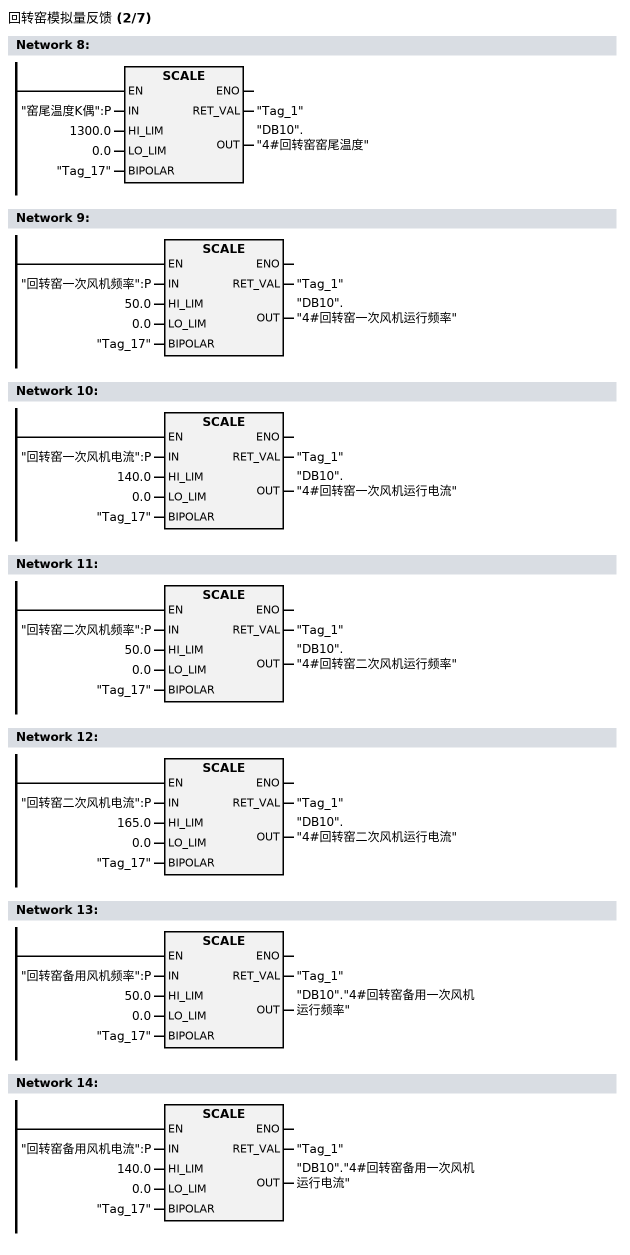
   "Tag_1" := SCALE(IN := "窑尾温度K偶":P,
                    HI_LIM := 1300.0,
                    LO_LIM := 0.0,
                    BIPOLAR := "Tag_17",
                    OUT => "DB10"."4#回转窑窑尾温度");
END_REGION

REGION Network 9
   "Tag_1" := SCALE(IN := "回转窑一次风机频率":P,
                    HI_LIM := 50.0,
                    LO_LIM := 0.0,
                    BIPOLAR := "Tag_17",
                    OUT => "DB10"."4#回转窑一次风机运行频率");
END_REGION

REGION Network 10
   "Tag_1" := SCALE(IN := "回转窑一次风机电流":P,
                    HI_LIM := 140.0,
                    LO_LIM := 0.0,
                    BIPOLAR := "Tag_17",
                    OUT => "DB10"."4#回转窑一次风机运行电流");
END_REGION

REGION Network 11
   "Tag_1" := SCALE(IN := "回转窑二次风机频率":P,
                    HI_LIM := 50.0,
                    LO_LIM := 0.0,
                    BIPOLAR := "Tag_17",
                    OUT => "DB10"."4#回转窑二次风机运行频率");
END_REGION

REGION Network 12
   "Tag_1" := SCALE(IN := "回转窑二次风机电流":P,
                    HI_LIM := 165.0,
                    LO_LIM := 0.0,
                    BIPOLAR := "Tag_17",
                    OUT => "DB10"."4#回转窑二次风机运行电流");
END_REGION

REGION Network 13
   "Tag_1" := SCALE(IN := "回转窑备用风机频率":P,
                    HI_LIM := 50.0,
                    LO_LIM := 0.0,
                    BIPOLAR := "Tag_17",
                    OUT => "DB10"."4#回转窑备用一次风机运行频率");
END_REGION

REGION Network 14
   "Tag_1" := SCALE(IN := "回转窑备用风机电流":P,
                    HI_LIM := 140.0,
                    LO_LIM := 0.0,
                    BIPOLAR := "Tag_17",
                    OUT => "DB10"."4#回转窑备用一次风机运行电流");
END_REGION

REGION Network 15
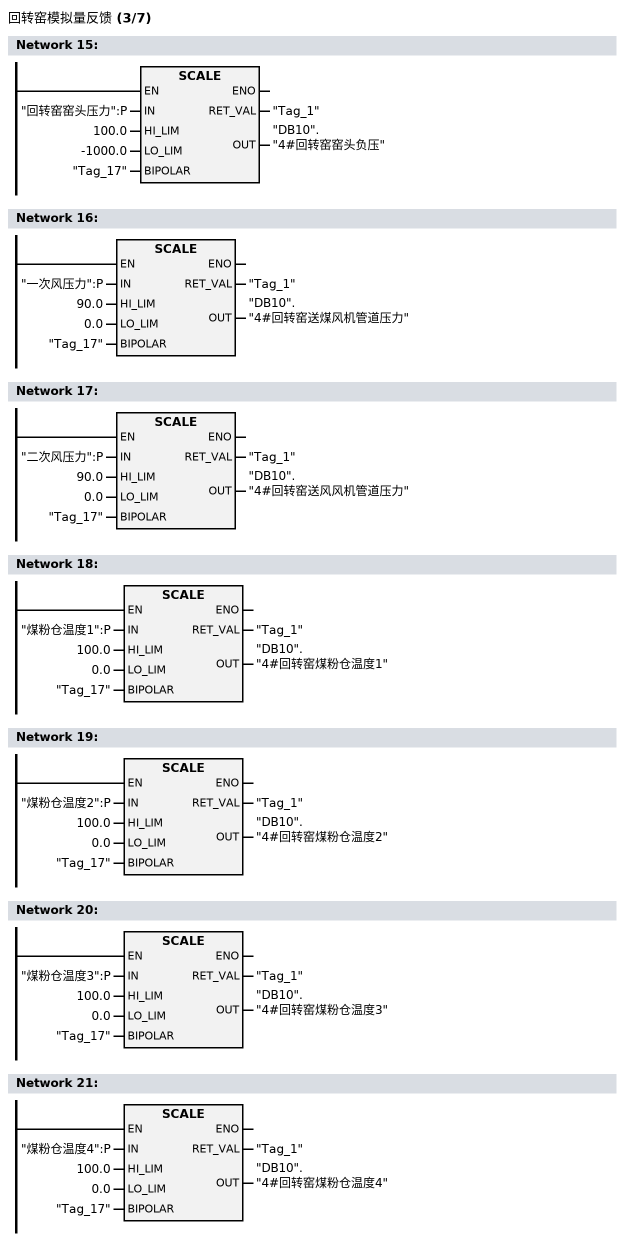
   "Tag_1" := SCALE(IN := "回转窑窑头压力":P,
                    HI_LIM := 100.0,
                    LO_LIM := -1000.0,
                    BIPOLAR := "Tag_17",
                    OUT => "DB10"."4#回转窑窑头负压");
END_REGION

REGION Network 16
   "Tag_1" := SCALE(IN := "一次风压力":P,
                    HI_LIM := 90.0,
                    LO_LIM := 0.0,
                    BIPOLAR := "Tag_17",
                    OUT => "DB10"."4#回转窑送煤风机管道压力");
END_REGION

REGION Network 17
   "Tag_1" := SCALE(IN := "二次风压力":P,
                    HI_LIM := 90.0,
                    LO_LIM := 0.0,
                    BIPOLAR := "Tag_17",
                    OUT => "DB10"."4#回转窑送风风机管道压力");
END_REGION

REGION Network 18
   "Tag_1" := SCALE(IN := "煤粉仓温度1":P,
                    HI_LIM := 100.0,
                    LO_LIM := 0.0,
                    BIPOLAR := "Tag_17",
                    OUT => "DB10"."4#回转窑煤粉仓温度1");
END_REGION

REGION Network 19
   "Tag_1" := SCALE(IN := "煤粉仓温度2":P,
                    HI_LIM := 100.0,
                    LO_LIM := 0.0,
                    BIPOLAR := "Tag_17",
                    OUT => "DB10"."4#回转窑煤粉仓温度2");
END_REGION

REGION Network 20
   "Tag_1" := SCALE(IN := "煤粉仓温度3":P,
                    HI_LIM := 100.0,
                    LO_LIM := 0.0,
                    BIPOLAR := "Tag_17",
                    OUT => "DB10"."4#回转窑煤粉仓温度3");
END_REGION

REGION Network 21
   "Tag_1" := SCALE(IN := "煤粉仓温度4":P,
                    HI_LIM := 100.0,
                    LO_LIM := 0.0,
                    BIPOLAR := "Tag_17",
                    OUT => "DB10"."4#回转窑煤粉仓温度4");
END_REGION

REGION Network 22
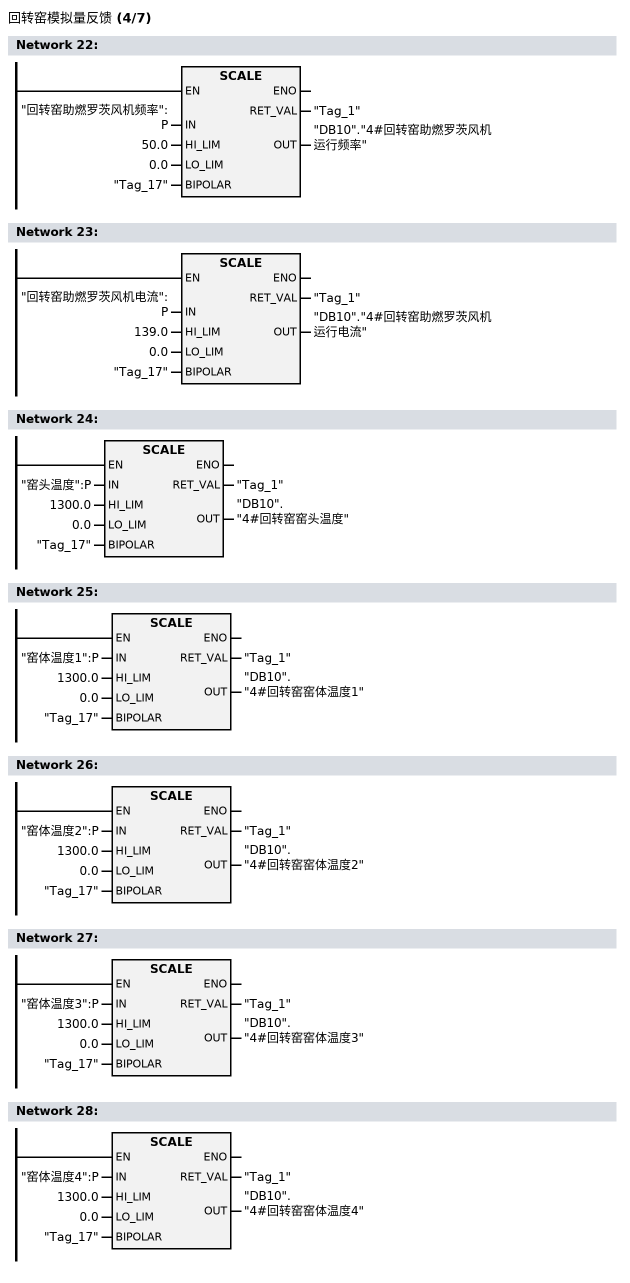
   "Tag_1" := SCALE(IN := "回转窑助燃罗茨风机频率":P,
                    HI_LIM := 50.0,
                    LO_LIM := 0.0,
                    BIPOLAR := "Tag_17",
                    OUT => "DB10"."4#回转窑助燃罗茨风机运行频率");
END_REGION

REGION Network 23
   "Tag_1" := SCALE(IN := "回转窑助燃罗茨风机电流":P,
                    HI_LIM := 139.0,
                    LO_LIM := 0.0,
                    BIPOLAR := "Tag_17",
                    OUT => "DB10"."4#回转窑助燃罗茨风机运行电流");
END_REGION

REGION Network 24
   "Tag_1" := SCALE(IN := "窑头温度":P,
                    HI_LIM := 1300.0,
                    LO_LIM := 0.0,
                    BIPOLAR := "Tag_17",
                    OUT => "DB10"."4#回转窑窑头温度");
END_REGION

REGION Network 25
   "Tag_1" := SCALE(IN := "窑体温度1":P,
                    HI_LIM := 1300.0,
                    LO_LIM := 0.0,
                    BIPOLAR := "Tag_17",
                    OUT => "DB10"."4#回转窑窑体温度1");
END_REGION

REGION Network 26
   "Tag_1" := SCALE(IN := "窑体温度2":P,
                    HI_LIM := 1300.0,
                    LO_LIM := 0.0,
                    BIPOLAR := "Tag_17",
                    OUT => "DB10"."4#回转窑窑体温度2");
END_REGION

REGION Network 27
   "Tag_1" := SCALE(IN := "窑体温度3":P,
                    HI_LIM := 1300.0,
                    LO_LIM := 0.0,
                    BIPOLAR := "Tag_17",
                    OUT => "DB10"."4#回转窑窑体温度3");
END_REGION

REGION Network 28
   "Tag_1" := SCALE(IN := "窑体温度4":P,
                    HI_LIM := 1300.0,
                    LO_LIM := 0.0,
                    BIPOLAR := "Tag_17",
                    OUT => "DB10"."4#回转窑窑体温度4");
END_REGION

REGION Network 29
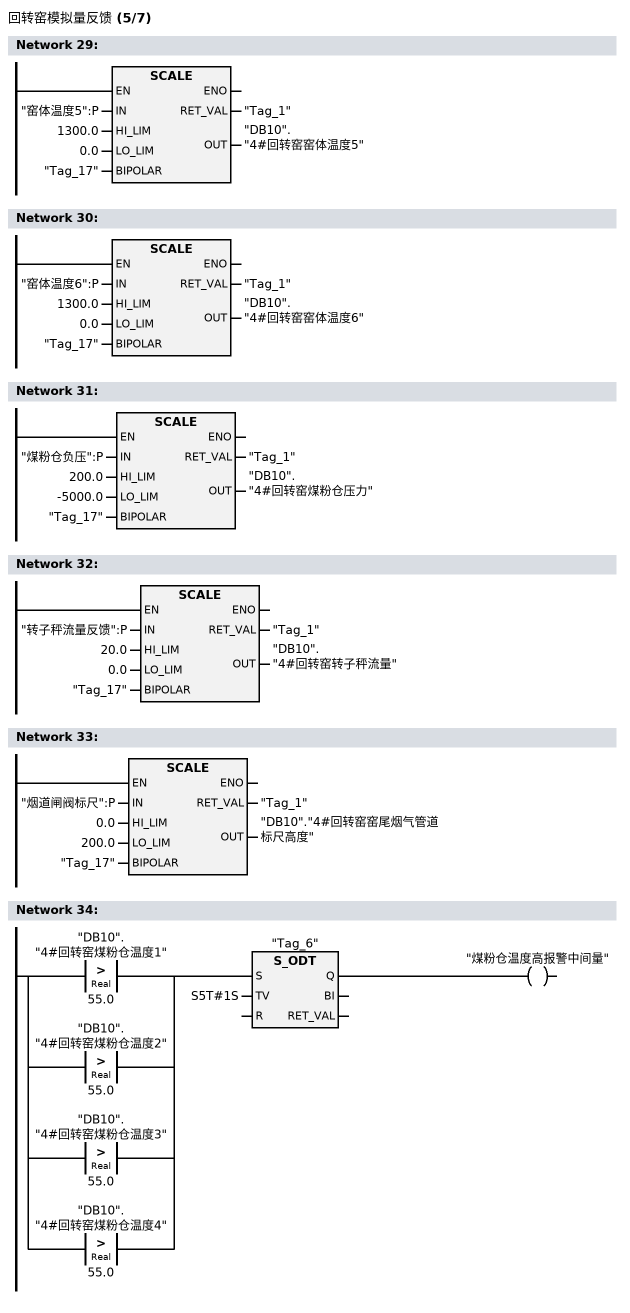
   "Tag_1" := SCALE(IN := "窑体温度5":P,
                    HI_LIM := 1300.0,
                    LO_LIM := 0.0,
                    BIPOLAR := "Tag_17",
                    OUT => "DB10"."4#回转窑窑体温度5");
END_REGION

REGION Network 30
   "Tag_1" := SCALE(IN := "窑体温度6":P,
                    HI_LIM := 1300.0,
                    LO_LIM := 0.0,
                    BIPOLAR := "Tag_17",
                    OUT => "DB10"."4#回转窑窑体温度6");
END_REGION

REGION Network 31
   "Tag_1" := SCALE(IN := "煤粉仓负压":P,
                    HI_LIM := 200.0,
                    LO_LIM := -5000.0,
                    BIPOLAR := "Tag_17",
                    OUT => "DB10"."4#回转窑煤粉仓压力");
END_REGION

REGION Network 32
   "Tag_1" := SCALE(IN := "转子秤流量反馈":P,
                    HI_LIM := 20.0,
                    LO_LIM := 0.0,
                    BIPOLAR := "Tag_17",
                    OUT => "DB10"."4#回转窑转子秤流量");
END_REGION

REGION Network 33
   "Tag_1" := SCALE(IN := "烟道闸阀标尺":P,
                    HI_LIM := 0.0,
                    LO_LIM := 200.0,
                    BIPOLAR := "Tag_17",
                    OUT => "DB10"."4#回转窑窑尾烟气管道标尺高度");
END_REGION

REGION Network 34
   RUNG wire#powerrail
      { S7_Templates := "SrcType := Real" } GT_Contact(in1 := "DB10"."4#回转窑煤粉仓温度1", in2 := 55.0)
      wire#w1
      S_ODT(T_NO := "Tag_6", TV := S5T#1S, R :=, BI =>, RET_VAL =>)
      Coil( "煤粉仓温度高报警中间量" )
   END_RUNG
   RUNG wire#powerrail
      { S7_Templates := "SrcType := Real" } GT_Contact(in1 := "DB10"."4#回转窑煤粉仓温度2", in2 := 55.0)
   END_RUNG wire#w1
   RUNG wire#powerrail
      { S7_Templates := "SrcType := Real" } GT_Contact(in1 := "DB10"."4#回转窑煤粉仓温度3", in2 := 55.0)
   END_RUNG wire#w1
   RUNG wire#powerrail
      { S7_Templates := "SrcType := Real" } GT_Contact(in1 := "DB10"."4#回转窑煤粉仓温度4", in2 := 55.0)
   END_RUNG wire#w1
   // the same network as SCL:
   #_s5time1 := S_ODT(T_NO := "Tag_6",
                      S := ("DB10"."4#回转窑煤粉仓温度1" > 55.0) OR ("DB10"."4#回转窑煤粉仓温度2" > 55.0) OR ("DB10"."4#回转窑煤粉仓温度3" > 55.0) OR ("DB10"."4#回转窑煤粉仓温度4" > 55.0),
                      TV := S5T#1S,
                      Q => #_w1);
   "煤粉仓温度高报警中间量" := #_w1;
END_REGION

REGION Network 35
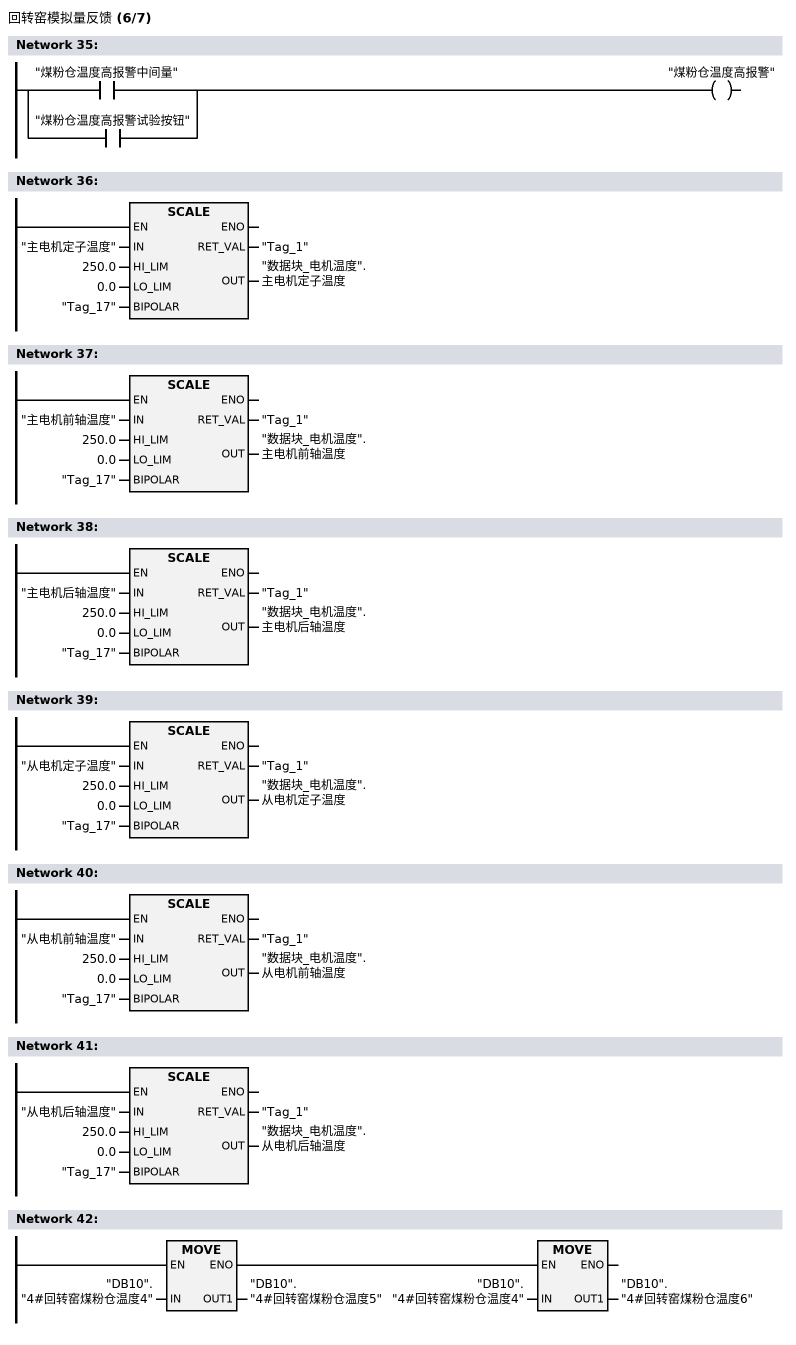
   RUNG wire#powerrail
      Contact( "煤粉仓温度高报警中间量" )
      wire#w1
      Coil( "煤粉仓温度高报警" )
   END_RUNG
   RUNG wire#powerrail
      Contact( "煤粉仓温度高报警试验按钮" )
   END_RUNG wire#w1
   // the same network as SCL:
   "煤粉仓温度高报警" := "煤粉仓温度高报警中间量" OR "煤粉仓温度高报警试验按钮";
END_REGION

REGION Network 36
   "Tag_1" := SCALE(IN := "主电机定子温度",
                    HI_LIM := 250.0,
                    LO_LIM := 0.0,
                    BIPOLAR := "Tag_17",
                    OUT => "数据块_电机温度".主电机定子温度);
END_REGION

REGION Network 37
   "Tag_1" := SCALE(IN := "主电机前轴温度",
                    HI_LIM := 250.0,
                    LO_LIM := 0.0,
                    BIPOLAR := "Tag_17",
                    OUT => "数据块_电机温度".主电机前轴温度);
END_REGION

REGION Network 38
   "Tag_1" := SCALE(IN := "主电机后轴温度",
                    HI_LIM := 250.0,
                    LO_LIM := 0.0,
                    BIPOLAR := "Tag_17",
                    OUT => "数据块_电机温度".主电机后轴温度);
END_REGION

REGION Network 39
   "Tag_1" := SCALE(IN := "从电机定子温度",
                    HI_LIM := 250.0,
                    LO_LIM := 0.0,
                    BIPOLAR := "Tag_17",
                    OUT => "数据块_电机温度".从电机定子温度);
END_REGION

REGION Network 40
   "Tag_1" := SCALE(IN := "从电机前轴温度",
                    HI_LIM := 250.0,
                    LO_LIM := 0.0,
                    BIPOLAR := "Tag_17",
                    OUT => "数据块_电机温度".从电机前轴温度);
END_REGION

REGION Network 41
   "Tag_1" := SCALE(IN := "从电机后轴温度",
                    HI_LIM := 250.0,
                    LO_LIM := 0.0,
                    BIPOLAR := "Tag_17",
                    OUT => "数据块_电机温度".从电机后轴温度);
END_REGION

REGION Network 42
   RUNG wire#powerrail
      Move(in := "DB10"."4#回转窑煤粉仓温度4", out1 => "DB10"."4#回转窑煤粉仓温度5")
      Move(in := "DB10"."4#回转窑煤粉仓温度4", out1 => "DB10"."4#回转窑煤粉仓温度6")
   END_RUNG
   // the same network as SCL:
   "DB10"."4#回转窑煤粉仓温度5" := "DB10"."4#回转窑煤粉仓温度4";
   "DB10"."4#回转窑煤粉仓温度6" := "DB10"."4#回转窑煤粉仓温度4";
END_REGION

REGION Network 43
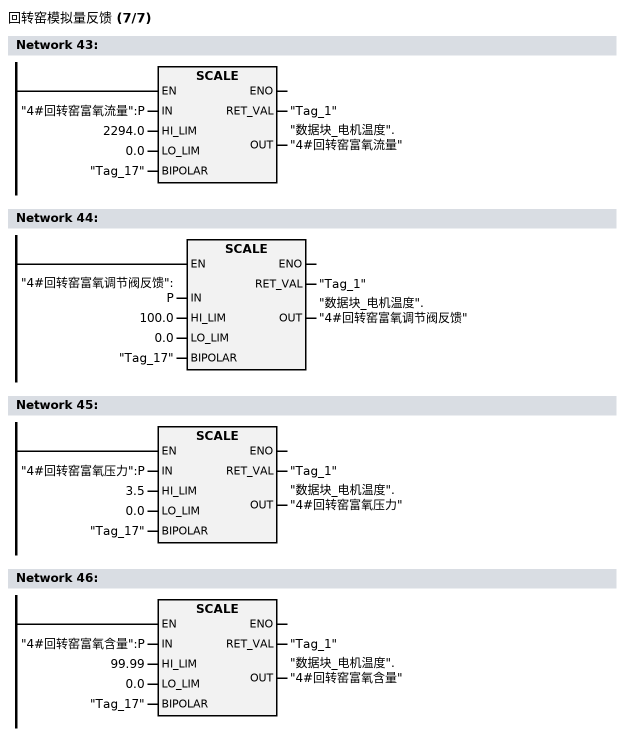
   "Tag_1" := SCALE(IN := "4#回转窑富氧流量":P,
                    HI_LIM := 2294.0,
                    LO_LIM := 0.0,
                    BIPOLAR := "Tag_17",
                    OUT => "数据块_电机温度"."4#回转窑富氧流量");
END_REGION

REGION Network 44
   "Tag_1" := SCALE(IN := "4#回转窑富氧调节阀反馈":P,
                    HI_LIM := 100.0,
                    LO_LIM := 0.0,
                    BIPOLAR := "Tag_17",
                    OUT => "数据块_电机温度"."4#回转窑富氧调节阀反馈");
END_REGION

REGION Network 45
   "Tag_1" := SCALE(IN := "4#回转窑富氧压力":P,
                    HI_LIM := 3.5,
                    LO_LIM := 0.0,
                    BIPOLAR := "Tag_17",
                    OUT => "数据块_电机温度"."4#回转窑富氧压力");
END_REGION

REGION Network 46
   "Tag_1" := SCALE(IN := "4#回转窑富氧含量":P,
                    HI_LIM := 99.99,
                    LO_LIM := 0.0,
                    BIPOLAR := "Tag_17",
                    OUT => "数据块_电机温度"."4#回转窑富氧含量");
END_REGION
END_FUNCTION

FUNCTION "回转窑风机控制" : Void   // FC13, LAD
{ S7_Optimized_Access := 'FALSE' }
VERSION : 0.1
   VAR_TEMP   // added for the SCL form of the ladder/FBD networks
      _w1 : Bool;
      _s5time1 : S5Time;
   END_VAR
BEGIN

REGION Network 1
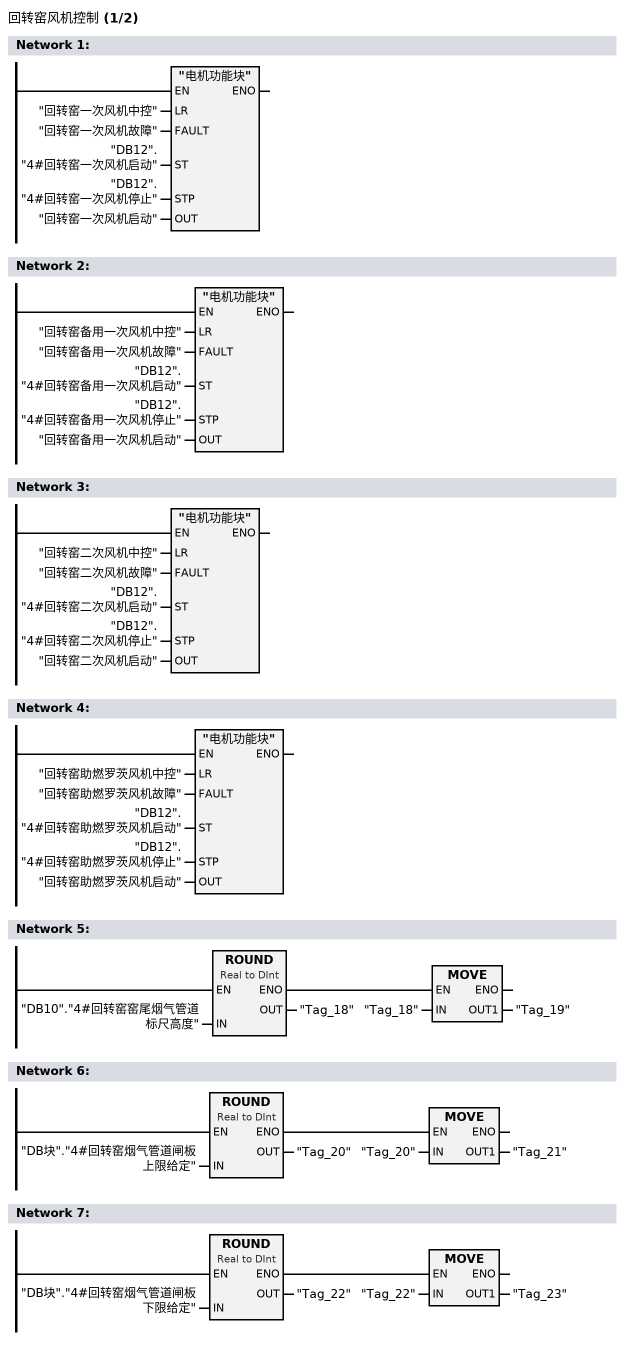
   RUNG wire#powerrail
      "电机功能块"(LR := "回转窑一次风机中控", FAULT := "回转窑一次风机故障", ST := "DB12"."4#回转窑一次风机启动", STP := "DB12"."4#回转窑一次风机停止", OUT := "回转窑一次风机启动")
   END_RUNG
   // the same network as SCL:
   "电机功能块"(LR := "回转窑一次风机中控",
           FAULT := "回转窑一次风机故障",
           ST := "DB12"."4#回转窑一次风机启动",
           STP := "DB12"."4#回转窑一次风机停止",
           OUT := "回转窑一次风机启动");
END_REGION

REGION Network 2
   RUNG wire#powerrail
      "电机功能块"(LR := "回转窑备用一次风机中控", FAULT := "回转窑备用一次风机故障", ST := "DB12"."4#回转窑备用一次风机启动", STP := "DB12"."4#回转窑备用一次风机停止", OUT := "回转窑备用一次风机启动")
   END_RUNG
   // the same network as SCL:
   "电机功能块"(LR := "回转窑备用一次风机中控",
           FAULT := "回转窑备用一次风机故障",
           ST := "DB12"."4#回转窑备用一次风机启动",
           STP := "DB12"."4#回转窑备用一次风机停止",
           OUT := "回转窑备用一次风机启动");
END_REGION

REGION Network 3
   RUNG wire#powerrail
      "电机功能块"(LR := "回转窑二次风机中控", FAULT := "回转窑二次风机故障", ST := "DB12"."4#回转窑二次风机启动", STP := "DB12"."4#回转窑二次风机停止", OUT := "回转窑二次风机启动")
   END_RUNG
   // the same network as SCL:
   "电机功能块"(LR := "回转窑二次风机中控",
           FAULT := "回转窑二次风机故障",
           ST := "DB12"."4#回转窑二次风机启动",
           STP := "DB12"."4#回转窑二次风机停止",
           OUT := "回转窑二次风机启动");
END_REGION

REGION Network 4
   RUNG wire#powerrail
      "电机功能块"(LR := "回转窑助燃罗茨风机中控", FAULT := "回转窑助燃罗茨风机故障", ST := "DB12"."4#回转窑助燃罗茨风机启动", STP := "DB12"."4#回转窑助燃罗茨风机停止", OUT := "回转窑助燃罗茨风机启动")
   END_RUNG
   // the same network as SCL:
   "电机功能块"(LR := "回转窑助燃罗茨风机中控",
           FAULT := "回转窑助燃罗茨风机故障",
           ST := "DB12"."4#回转窑助燃罗茨风机启动",
           STP := "DB12"."4#回转窑助燃罗茨风机停止",
           OUT := "回转窑助燃罗茨风机启动");
END_REGION

REGION Network 5
   RUNG wire#powerrail
      { S7_Templates := "[SrcType := Real, DestType := DInt]"; S7_GenerateENO := "TRUE" } Round(in := "DB10"."4#回转窑窑尾烟气管道标尺高度", out => "Tag_18")
      { S7_GenerateENO := "TRUE" } Move(in := "Tag_18", out1 => "Tag_19")
   END_RUNG
   // the same network as SCL:
   // ENO of a box is taken as its EN; it also drops when the box reports an error
   "Tag_18" := ROUND("DB10"."4#回转窑窑尾烟气管道标尺高度");
   "Tag_19" := "Tag_18";
END_REGION

REGION Network 6
   RUNG wire#powerrail
      { S7_Templates := "[SrcType := Real, DestType := DInt]"; S7_GenerateENO := "TRUE" } Round(in := "DB块"."4#回转窑烟气管道闸板上限给定", out => "Tag_20")
      { S7_GenerateENO := "TRUE" } Move(in := "Tag_20", out1 => "Tag_21")
   END_RUNG
   // the same network as SCL:
   // ENO of a box is taken as its EN; it also drops when the box reports an error
   "Tag_20" := ROUND("DB块"."4#回转窑烟气管道闸板上限给定");
   "Tag_21" := "Tag_20";
END_REGION

REGION Network 7
   RUNG wire#powerrail
      { S7_Templates := "[SrcType := Real, DestType := DInt]"; S7_GenerateENO := "TRUE" } Round(in := "DB块"."4#回转窑烟气管道闸板下限给定", out => "Tag_22")
      { S7_GenerateENO := "TRUE" } Move(in := "Tag_22", out1 => "Tag_23")
   END_RUNG
   // the same network as SCL:
   // ENO of a box is taken as its EN; it also drops when the box reports an error
   "Tag_22" := ROUND("DB块"."4#回转窑烟气管道闸板下限给定");
   "Tag_23" := "Tag_22";
END_REGION

REGION Network 8
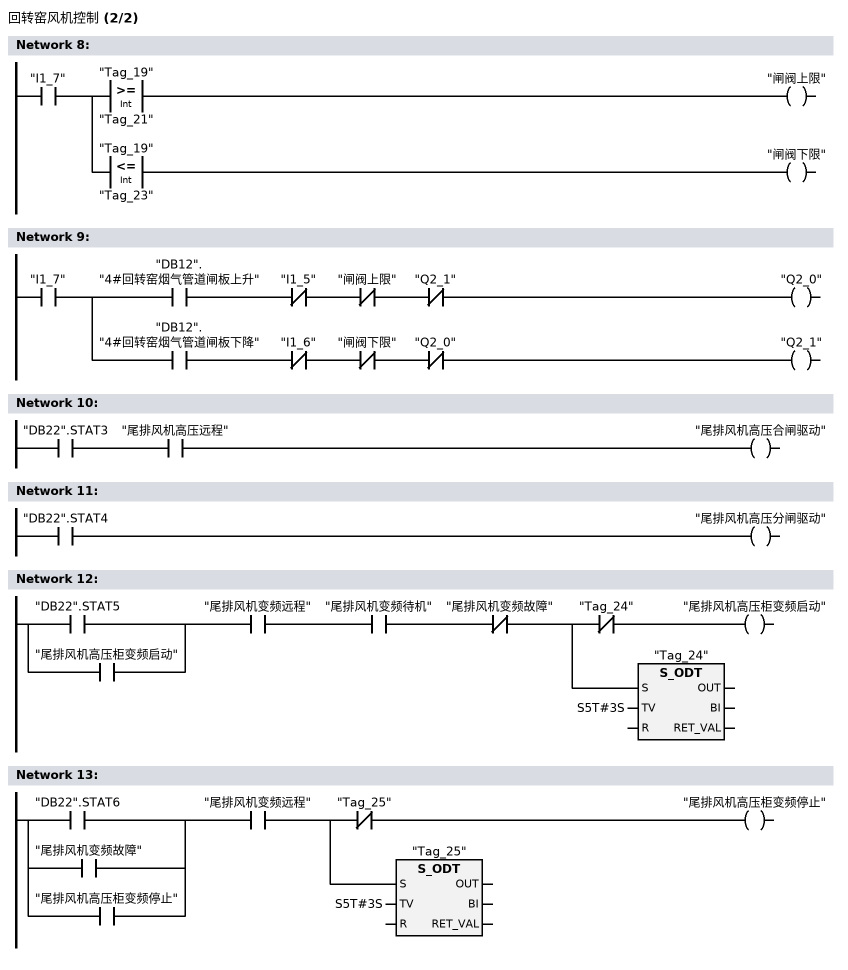
   RUNG wire#powerrail
      Contact( "I1_7" )
      wire#w1
      { S7_Templates := "SrcType := Int" } GE_Contact(in1 := "Tag_19", in2 := "Tag_21")
      Coil( "闸阀上限" )
   END_RUNG
   RUNG wire#w1
      { S7_Templates := "SrcType := Int" } LE_Contact(in1 := "Tag_19", in2 := "Tag_23")
      Coil( "闸阀下限" )
   END_RUNG
   // the same network as SCL:
   "闸阀上限" := "I1_7" AND ("Tag_19" >= "Tag_21");
   "闸阀下限" := "I1_7" AND ("Tag_19" <= "Tag_23");
END_REGION

REGION Network 9
   RUNG wire#powerrail
      Contact( "I1_7" )
      wire#w1
      Contact( "DB12"."4#回转窑烟气管道闸板上升" )
      I_Contact( "I1_5" )
      I_Contact( "闸阀上限" )
      I_Contact( "Q2_1" )
      Coil( "Q2_0" )
   END_RUNG
   RUNG wire#w1
      Contact( "DB12"."4#回转窑烟气管道闸板下降" )
      I_Contact( "I1_6" )
      I_Contact( "闸阀下限" )
      I_Contact( "Q2_0" )
      Coil( "Q2_1" )
   END_RUNG
   // the same network as SCL:
   "Q2_0" := "I1_7" AND "DB12"."4#回转窑烟气管道闸板上升" AND NOT "I1_5" AND NOT "闸阀上限" AND NOT "Q2_1";
   "Q2_1" := "I1_7" AND "DB12"."4#回转窑烟气管道闸板下降" AND NOT "I1_6" AND NOT "闸阀下限" AND NOT "Q2_0";
END_REGION

REGION Network 10
   RUNG wire#powerrail
      Contact( "DB22".STAT3 )
      Contact( "尾排风机高压远程" )
      Coil( "尾排风机高压合闸驱动" )
   END_RUNG
   // the same network as SCL:
   "尾排风机高压合闸驱动" := "DB22".STAT3 AND "尾排风机高压远程";
END_REGION

REGION Network 11
   RUNG wire#powerrail
      Contact( "DB22".STAT4 )
      Coil( "尾排风机高压分闸驱动" )
   END_RUNG
   // the same network as SCL:
   "尾排风机高压分闸驱动" := "DB22".STAT4;
END_REGION

REGION Network 12
   RUNG wire#powerrail
      Contact( "DB22".STAT5 )
      wire#w1
      Contact( "尾排风机变频远程" )
      Contact( "尾排风机变频待机" )
      I_Contact( "尾排风机变频故障" )
      wire#w2
      I_Contact( "Tag_24" )
      Coil( "尾排风机高压柜变频启动" )
   END_RUNG
   RUNG wire#powerrail
      Contact( "尾排风机高压柜变频启动" )
   END_RUNG wire#w1
   RUNG wire#w2
      S_ODT(T_NO := "Tag_24", TV := S5T#3S, R :=, BI =>, RET_VAL =>)
   END_RUNG
   // the same network as SCL:
   #_w1 := ("DB22".STAT5 OR "尾排风机高压柜变频启动") AND "尾排风机变频远程" AND "尾排风机变频待机" AND NOT "尾排风机变频故障";
   "尾排风机高压柜变频启动" := #_w1 AND NOT "Tag_24";
   #_s5time1 := S_ODT(T_NO := "Tag_24", S := #_w1, TV := S5T#3S);
END_REGION

REGION Network 13
   RUNG wire#powerrail
      Contact( "DB22".STAT6 )
      wire#w1
      Contact( "尾排风机变频远程" )
      wire#w2
      I_Contact( "Tag_25" )
      Coil( "尾排风机高压柜变频停止" )
   END_RUNG
   RUNG wire#powerrail
      Contact( "尾排风机变频故障" )
   END_RUNG wire#w1
   RUNG wire#powerrail
      Contact( "尾排风机高压柜变频停止" )
   END_RUNG wire#w1
   RUNG wire#w2
      S_ODT(T_NO := "Tag_25", TV := S5T#3S, R :=, BI =>, RET_VAL =>)
   END_RUNG
   // the same network as SCL:
   #_w1 := ("DB22".STAT6 OR "尾排风机变频故障" OR "尾排风机高压柜变频停止") AND "尾排风机变频远程";
   "尾排风机高压柜变频停止" := #_w1 AND NOT "Tag_25";
   #_s5time1 := S_ODT(T_NO := "Tag_25", S := #_w1, TV := S5T#3S);
END_REGION
END_FUNCTION

FUNCTION "回转窑模拟量给定" : Void   // FC14, LAD
{ S7_Optimized_Access := 'FALSE' }
VERSION : 0.1
BEGIN

REGION Network 1
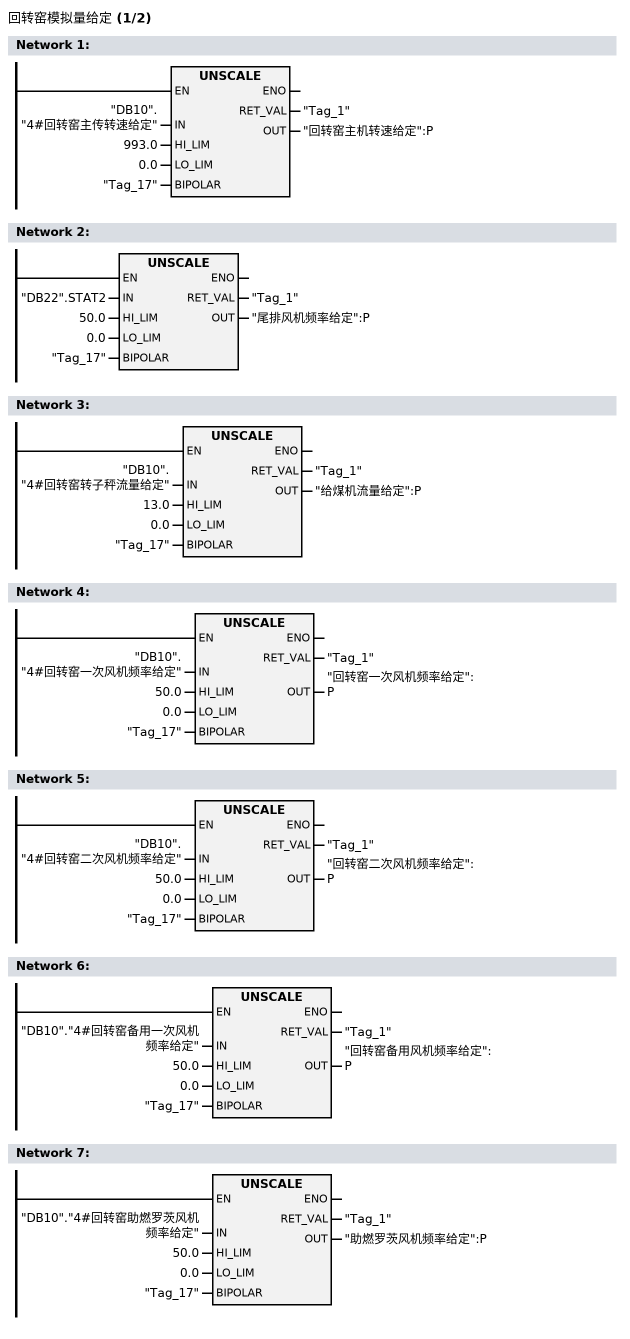
   "Tag_1" := UNSCALE(IN := "DB10"."4#回转窑主传转速给定",
                      HI_LIM := 993.0,
                      LO_LIM := 0.0,
                      BIPOLAR := "Tag_17",
                      OUT => "回转窑主机转速给定":P);
END_REGION

REGION Network 2
   "Tag_1" := UNSCALE(IN := "DB22".STAT2,
                      HI_LIM := 50.0,
                      LO_LIM := 0.0,
                      BIPOLAR := "Tag_17",
                      OUT => "尾排风机频率给定":P);
END_REGION

REGION Network 3
   "Tag_1" := UNSCALE(IN := "DB10"."4#回转窑转子秤流量给定",
                      HI_LIM := 13.0,
                      LO_LIM := 0.0,
                      BIPOLAR := "Tag_17",
                      OUT => "给煤机流量给定":P);
END_REGION

REGION Network 4
   "Tag_1" := UNSCALE(IN := "DB10"."4#回转窑一次风机频率给定",
                      HI_LIM := 50.0,
                      LO_LIM := 0.0,
                      BIPOLAR := "Tag_17",
                      OUT => "回转窑一次风机频率给定":P);
END_REGION

REGION Network 5
   "Tag_1" := UNSCALE(IN := "DB10"."4#回转窑二次风机频率给定",
                      HI_LIM := 50.0,
                      LO_LIM := 0.0,
                      BIPOLAR := "Tag_17",
                      OUT => "回转窑二次风机频率给定":P);
END_REGION

REGION Network 6
   "Tag_1" := UNSCALE(IN := "DB10"."4#回转窑备用一次风机频率给定",
                      HI_LIM := 50.0,
                      LO_LIM := 0.0,
                      BIPOLAR := "Tag_17",
                      OUT => "回转窑备用风机频率给定":P);
END_REGION

REGION Network 7
   "Tag_1" := UNSCALE(IN := "DB10"."4#回转窑助燃罗茨风机频率给定",
                      HI_LIM := 50.0,
                      LO_LIM := 0.0,
                      BIPOLAR := "Tag_17",
                      OUT => "助燃罗茨风机频率给定":P);
END_REGION

REGION Network 8
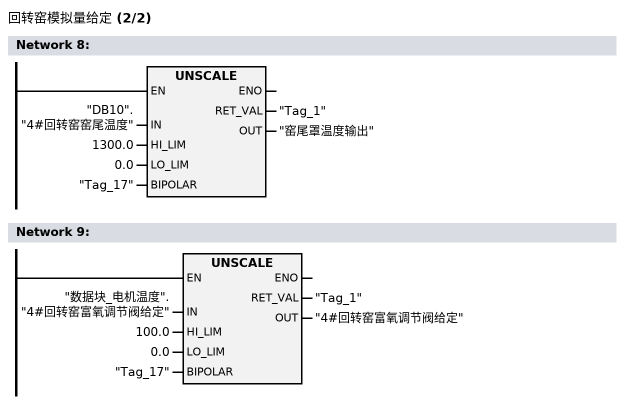
   "Tag_1" := UNSCALE(IN := "DB10"."4#回转窑窑尾温度",
                      HI_LIM := 1300.0,
                      LO_LIM := 0.0,
                      BIPOLAR := "Tag_17",
                      OUT => "窑尾罩温度输出");
END_REGION

REGION Network 9
   "Tag_1" := UNSCALE(IN := "数据块_电机温度"."4#回转窑富氧调节阀给定",
                      HI_LIM := 100.0,
                      LO_LIM := 0.0,
                      BIPOLAR := "Tag_17",
                      OUT => "4#回转窑富氧调节阀给定");
END_REGION
END_FUNCTION

FUNCTION "DP&MODBUS通讯" : Void   // FC15, LAD
{ S7_Optimized_Access := 'FALSE' }
VERSION : 0.1
BEGIN

REGION Network 1
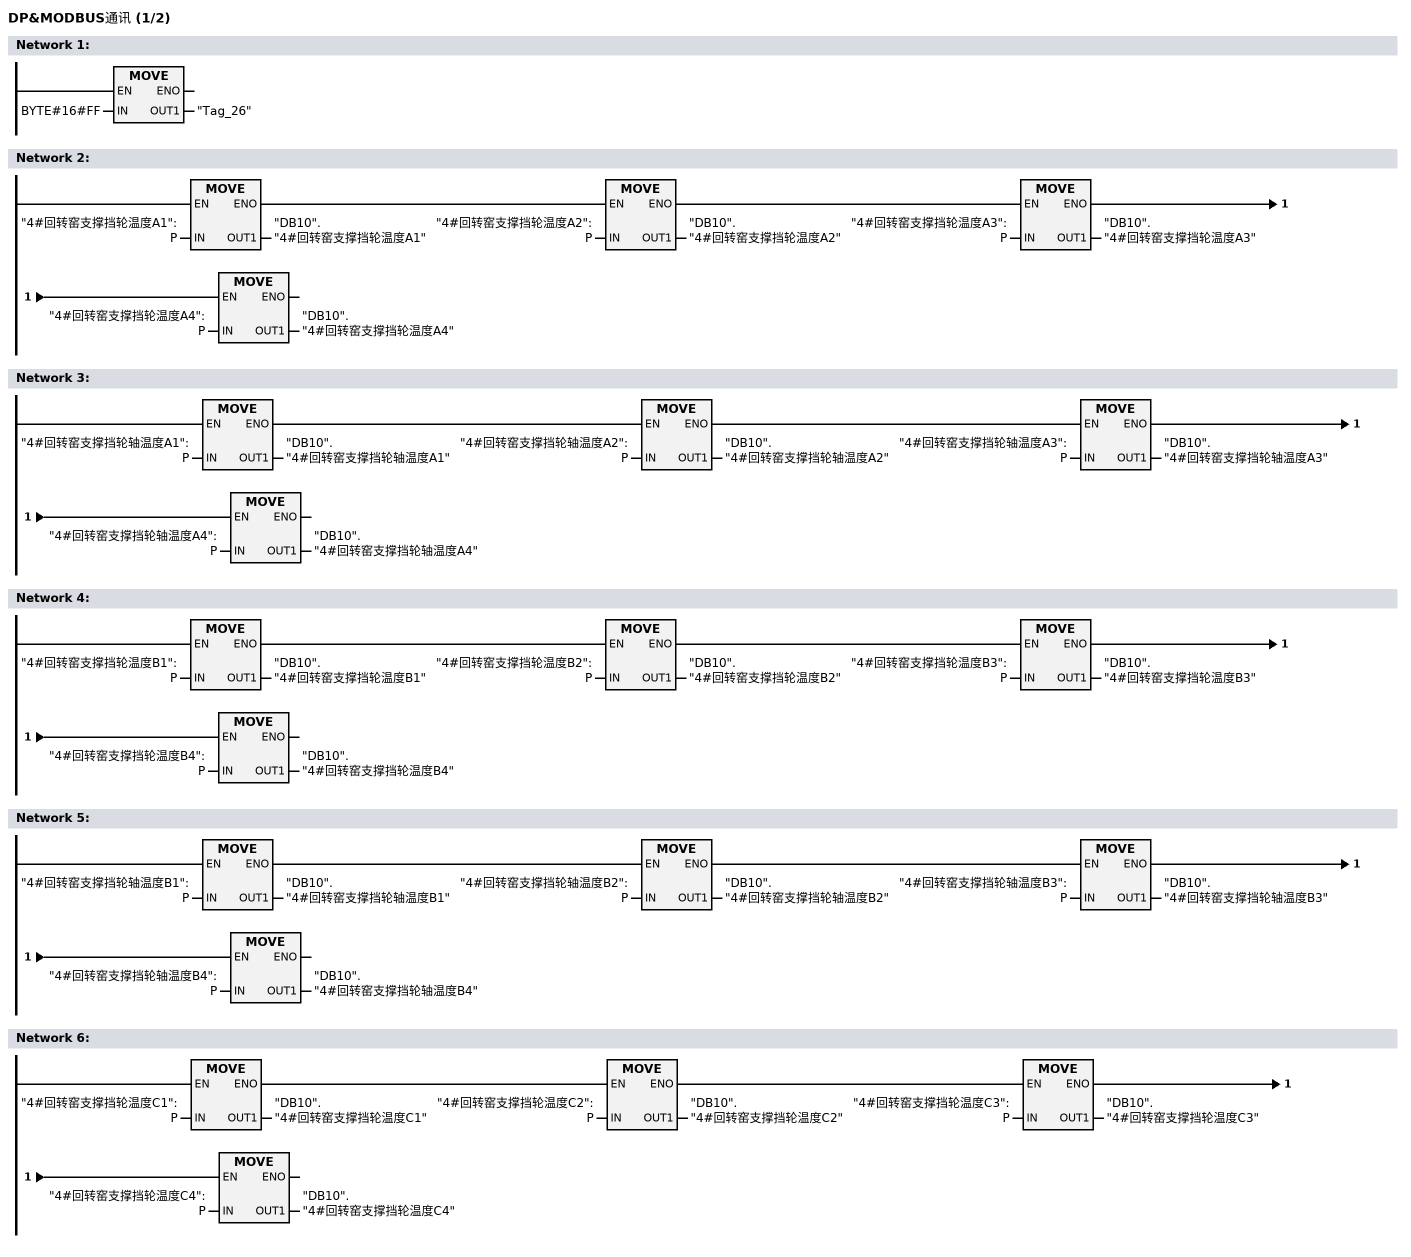
   RUNG wire#powerrail
      { S7_GenerateENO := "TRUE" } Move(in := BYTE#16#FF, out1 => "Tag_26")
   END_RUNG
   // the same network as SCL:
   "Tag_26" := BYTE#16#FF;
END_REGION

REGION Network 2
   RUNG wire#powerrail
      { S7_GenerateENO := "TRUE" } Move(in := "4#回转窑支撑挡轮温度A1":P, out1 => "DB10"."4#回转窑支撑挡轮温度A1")
      { S7_GenerateENO := "TRUE" } Move(in := "4#回转窑支撑挡轮温度A2":P, out1 => "DB10"."4#回转窑支撑挡轮温度A2")
      { S7_GenerateENO := "TRUE" } Move(in := "4#回转窑支撑挡轮温度A3":P, out1 => "DB10"."4#回转窑支撑挡轮温度A3")
      { S7_GenerateENO := "TRUE" } Move(in := "4#回转窑支撑挡轮温度A4":P, out1 => "DB10"."4#回转窑支撑挡轮温度A4")
   END_RUNG
   // the same network as SCL:
   // ENO of a box is taken as its EN; it also drops when the box reports an error
   "DB10"."4#回转窑支撑挡轮温度A1" := "4#回转窑支撑挡轮温度A1":P;
   "DB10"."4#回转窑支撑挡轮温度A2" := "4#回转窑支撑挡轮温度A2":P;
   "DB10"."4#回转窑支撑挡轮温度A3" := "4#回转窑支撑挡轮温度A3":P;
   "DB10"."4#回转窑支撑挡轮温度A4" := "4#回转窑支撑挡轮温度A4":P;
END_REGION

REGION Network 3
   RUNG wire#powerrail
      { S7_GenerateENO := "TRUE" } Move(in := "4#回转窑支撑挡轮轴温度A1":P, out1 => "DB10"."4#回转窑支撑挡轮轴温度A1")
      { S7_GenerateENO := "TRUE" } Move(in := "4#回转窑支撑挡轮轴温度A2":P, out1 => "DB10"."4#回转窑支撑挡轮轴温度A2")
      { S7_GenerateENO := "TRUE" } Move(in := "4#回转窑支撑挡轮轴温度A3":P, out1 => "DB10"."4#回转窑支撑挡轮轴温度A3")
      { S7_GenerateENO := "TRUE" } Move(in := "4#回转窑支撑挡轮轴温度A4":P, out1 => "DB10"."4#回转窑支撑挡轮轴温度A4")
   END_RUNG
   // the same network as SCL:
   // ENO of a box is taken as its EN; it also drops when the box reports an error
   "DB10"."4#回转窑支撑挡轮轴温度A1" := "4#回转窑支撑挡轮轴温度A1":P;
   "DB10"."4#回转窑支撑挡轮轴温度A2" := "4#回转窑支撑挡轮轴温度A2":P;
   "DB10"."4#回转窑支撑挡轮轴温度A3" := "4#回转窑支撑挡轮轴温度A3":P;
   "DB10"."4#回转窑支撑挡轮轴温度A4" := "4#回转窑支撑挡轮轴温度A4":P;
END_REGION

REGION Network 4
   RUNG wire#powerrail
      { S7_GenerateENO := "TRUE" } Move(in := "4#回转窑支撑挡轮温度B1":P, out1 => "DB10"."4#回转窑支撑挡轮温度B1")
      { S7_GenerateENO := "TRUE" } Move(in := "4#回转窑支撑挡轮温度B2":P, out1 => "DB10"."4#回转窑支撑挡轮温度B2")
      { S7_GenerateENO := "TRUE" } Move(in := "4#回转窑支撑挡轮温度B3":P, out1 => "DB10"."4#回转窑支撑挡轮温度B3")
      { S7_GenerateENO := "TRUE" } Move(in := "4#回转窑支撑挡轮温度B4":P, out1 => "DB10"."4#回转窑支撑挡轮温度B4")
   END_RUNG
   // the same network as SCL:
   // ENO of a box is taken as its EN; it also drops when the box reports an error
   "DB10"."4#回转窑支撑挡轮温度B1" := "4#回转窑支撑挡轮温度B1":P;
   "DB10"."4#回转窑支撑挡轮温度B2" := "4#回转窑支撑挡轮温度B2":P;
   "DB10"."4#回转窑支撑挡轮温度B3" := "4#回转窑支撑挡轮温度B3":P;
   "DB10"."4#回转窑支撑挡轮温度B4" := "4#回转窑支撑挡轮温度B4":P;
END_REGION
